
screen "eProC - 08 Descargador" 1280x768, template "Template"
   Button "Botón_4" at 220,383 size 93x33; TextOff 'Avance'
      on Press: SetTag("DB_OP.RC2", 70); SetBit("DB_OP.OP_SELMANU2")
      Visibility <- "MANU"
      Appearance <- "DB_OP.RC2"
   Button "Botón_5" at 220,421 size 93x33; TextOff 'Retroceso'
      on Press: SetTag("DB_OP.RC2", 71); SetBit("DB_OP.OP_SELMANU2")
      Visibility <- "MANU"
      Appearance <- "DB_OP.RC2"
   TextField "Campo de texto_5" at 229,340 size 85x23; Text 'Descargador'
      Visibility <- "MANU"
   Rectangle "Rectángulo_1" at 204,336 size 131x136
      Visibility <- "MANU"
   GraphicIOField "Campo ES gráfico_7" at 384,79 size 557x426; PictureList "Grupo 3 - Descargador"
      ProcessValue <- "Alarma_Descargador"
   Polygon "Polígono_4" at 443,271 size 39x59
      Visibility <- "Descargador-PiezaPresente"
   Polygon "Polígono_3" at 442,238 size 206x167
      Visibility <- "Descargador-PiezaPresente"
   Circle "Cercle_3" at 740,408 size 12x12
      Appearance <- "31S3"
   Circle "Cercle_4" at 693,373 size 12x12
      Appearance <- "31S8"
   Circle "Cercle_5" at 488,408 size 12x12
      Appearance <- "26S2"
   TextField "Campo de texto_1" at 890,544 size 173x22; Text '31S3 - Descargador Atrás'
   TextField "Campo de texto_2" at 557,516 size 195x22; Text '31S2 - Descargador Adelante'
   TextField "Campo de texto_3" at 818,279 size 193x22; Text '31S8 - Pieza en Descargador'
   Circle "Cercle_6" at 464,388 size 12x12
      Appearance <- "36S12"
   TextField "Campo de texto_4" at 534,549 size 294x22; Text '36S12 - Descargador en Posición Intermedia'
   Polygon "Polígono_2" at 450,217 size 81x72
      Visibility <- "Descargador-PiezaPresente"
   Polygon "Polígono_5" at 506,64 size 228x201
      Visibility <- "Descargador-PiezaPresente"
   Polygon "Polígono_1" at 543,118 size 206x170
      Visibility <- "Descargador-PiezaPresente"
   Polygon "Polígono_7" at 631,109 size 118x70
      Visibility <- "Descargador-PiezaPresente"
   Polygon "Polígono_8" at 625,64 size 112x67
      Visibility <- "Descargador-PiezaPresente"
   Rectangle "Rectángulo_2" at 204,336 size 131x32
      Visibility <- "MANU"
   Button "Template_Plantilla_Botón_3" at 1,688 size 130x29; TextOff 'DESCARGADOR'
   Button "Plantilla_Botón_1" at 1,715 size 130x53; TextOff 'PRINCIPAL'
      on Click: ActivateScreen("eProC - Principal", 0)
   Button "Template_Plantilla_Bouton_2" at 1085,715 size 193x53; TextOff 'ALARMAS / DEFAUT'
      on Press: ActivateScreen("eProC - Alarmas", 0)
      Visibility <- "DB_OP.P_DEFAUT"

screen "Gesión de Usuarios" 1280x768, template "Template"
   UserView "Visor de usuarios_1" at 28,48 size 1215x366
   Button "Botón_1" at 1059,488 size 176x56; TextOff 'Cerrar Sesión'
      on Activate: function_f23ef4c9()
   Button "Template_Plantilla_Botón_2" at 573,715 size 70x53; TextOff 'Text'; PictureOn "Usuario"; PictureOff "Usuario"; Authorization "Nivel 2"
      on Activate: ActivateScreen("Gesión de Usuarios", 0)
   Button "Template_Plantilla_Bouton_2" at 1085,715 size 193x53; TextOff 'ALARMAS / DEFAUT'
      on Press: ActivateScreen("eProC - Alarmas", 0)
      Visibility <- "DB_OP.P_DEFAUT"

screen "eProC - Historal" 1280x768, template "Template"
   AlarmView "Visor de avisos_1" at 29,48 size 1218x605; AlarmLog "Fichero_de_avisos_1"
   Button "Template_Plantilla_Botón_3" at 1085,688 size 193x29; TextOff 'HISTORIAL'
   Button "Template_Plantilla_Bouton_0" at 1085,715 size 193x53; TextOff 'ALARMAS / DEFAUT'
      on Press: ActivateScreen("eProC - Alarmas", 0)
   Button "Template_Plantilla_Bouton_2" at 1085,715 size 193x53; TextOff 'ALARMAS / DEFAUT'
      on Press: ActivateScreen("eProC - Alarmas", 0)
      Visibility <- "DB_OP.P_DEFAUT"

screen "eProC - Diagnóstico" 1280x768, template "Template"
   SysDiagControl "Sistema Visor de diagnóstico_1" at 16,30 size 1246x670; InfoArea_RootNodeText 'PLC Roll Forming / Installation'; NavigationPath_RootText 'Diagnóstico de Hardware / Vue d'ensemble du diagnostic'; NavigationpathDiagbufferText 'Búfer de diagnóstico / Vue du tampon de diagnostic'

screen "eProC - Estampado Alm 1" 1280x768, template "Template"
   TextField "Campo de texto_14" at 18,45 size 97x28; Text 'Almacén 1'
   TextField "Campo de texto_2" at 283,429 size 97x22; Text 'Herramienta 2'
   TextField "Campo de texto_3" at 283,157 size 97x22; Text 'Herramienta 1'
   TextField "Campo de texto_1" at 733,81 size 25x28; Text 'F1'
   TextField "Campo de texto_4" at 573,81 size 25x28; Text 'F3'
   TextField "Campo de texto_5" at 733,338 size 25x28; Text 'F2'
   TextField "Campo de texto_6" at 573,338 size 25x28; Text 'F4'
   TextField "Campo de texto_7" at 468,652 size 324x28; Text 'Resolución Incremento/Decremento'
   Button "Botón_1" at 754,150 size 40x40; TextOff 'Text'; PictureOff "outline_arrow_forward_ios_white_18dp"
      on Click: SetTag("PL_Dec_F_A1", 1)
   Button "Botón_2" at 698,150 size 40x40; TextOff 'Text'; PictureOff "outline_arrow_back_ios_white_18dp"
      on Click: SetTag("PL_Inc_F_A1", 1)
   Button "Botón_3" at 594,150 size 40x40; TextOff 'Text'; PictureOff "outline_arrow_forward_ios_white_18dp"
      on Click: SetTag("PL_Dec_F_A1", 3)
   Button "Botón_4" at 538,150 size 40x40; TextOff 'Text'; PictureOff "outline_arrow_back_ios_white_18dp"
      on Click: SetTag("PL_Inc_F_A1", 3)
   Button "Botón_5" at 754,406 size 40x40; TextOff 'Text'; PictureOff "outline_arrow_forward_ios_white_18dp"
      on Click: SetTag("PL_Dec_F_A1", 2)
   Button "Botón_6" at 698,406 size 40x40; TextOff 'Text'; PictureOff "outline_arrow_back_ios_white_18dp"
      on Click: SetTag("PL_Inc_F_A1", 2)
   Button "Botón_7" at 594,406 size 40x40; TextOff 'Text'; PictureOff "outline_arrow_forward_ios_white_18dp"
      on Click: SetTag("PL_Dec_F_A1", 4)
   Button "Botón_8" at 538,406 size 40x40; TextOff 'Text'; PictureOff "outline_arrow_back_ios_white_18dp"
      on Click: SetTag("PL_Inc_F_A1", 4)
   GraphicView "Visor de gráficos_7" at 263,452 size 138x75; Picture "F1-3 EMR2"
   GraphicView "Visor de gráficos_8" at 263,517 size 138x75; Picture "F2-4 EMR2"
   GraphicView "Visor de gráficos_2" at 263,180 size 138x75; Picture "EMR2"
   GraphicView "Visor de gráficos_3" at 263,245 size 138x75; Picture "F1-3 EMR2"
   IOField "Campo ES_1" at 698,109 size 96x32; FormatPattern s999999
      ProcessValue <- "Almacén 1\PAlmacén.F1"
   IOField "Campo ES_2" at 536,109 size 96x32; FormatPattern s999999
      ProcessValue <- "Almacén 1\PAlmacén.F3"
   IOField "Campo ES_3" at 698,366 size 96x32; FormatPattern s999999
      ProcessValue <- "Almacén 1\PAlmacén.F2"
   IOField "Campo ES_4" at 536,366 size 96x32; FormatPattern s999999
      ProcessValue <- "Almacén 1\PAlmacén.F4"
   IOField "Campo ES_5" at 787,653 size 96x32; FormatPattern 999999
      ProcessValue <- "PL_Resoluc_INCDECF"
   IOField "Champ E/S_1" at 122,48 size 410x24; FormatPattern ????????????????????
      ProcessValue <- "Almacén 1\PAlmacén.Nombre"

screen "eProC - Estampado Alm 2" 1280x768, template "Template"
   TextField "Campo de texto_14" at 18,45 size 97x28; Text 'Almacén 2'
   TextField "Campo de texto_2" at 283,429 size 97x22; Text 'Herramienta 2'
   TextField "Campo de texto_3" at 283,157 size 97x22; Text 'Herramienta 1'
   TextField "Campo de texto_1" at 733,81 size 25x28; Text 'F1'
   TextField "Campo de texto_4" at 572,81 size 25x28; Text 'F3'
   TextField "Campo de texto_5" at 733,338 size 25x28; Text 'F2'
   TextField "Campo de texto_6" at 572,338 size 25x28; Text 'F4'
   TextField "Campo de texto_7" at 468,652 size 324x28; Text 'Resolución Incremento/Decremento'
   Button "Botón_1" at 754,150 size 40x40; TextOff 'Text'; PictureOff "outline_arrow_forward_ios_white_18dp"
      on Click: SetTag("PL_Dec_F_A2", 1)
   Button "Botón_2" at 698,150 size 40x40; TextOff 'Text'; PictureOff "outline_arrow_back_ios_white_18dp"
      on Click: SetTag("PL_Inc_F_A2", 1)
   Button "Botón_3" at 593,150 size 40x40; TextOff 'Text'; PictureOff "outline_arrow_forward_ios_white_18dp"
      on Click: SetTag("PL_Dec_F_A2", 3)
   Button "Botón_4" at 537,150 size 40x40; TextOff 'Text'; PictureOff "outline_arrow_back_ios_white_18dp"
      on Click: SetTag("PL_Inc_F_A2", 3)
   Button "Botón_5" at 754,406 size 40x40; TextOff 'Text'; PictureOff "outline_arrow_forward_ios_white_18dp"
      on Click: SetTag("PL_Dec_F_A2", 2)
   Button "Botón_6" at 698,406 size 40x40; TextOff 'Text'; PictureOff "outline_arrow_back_ios_white_18dp"
      on Click: SetTag("PL_Inc_F_A2", 2)
   Button "Botón_7" at 593,406 size 40x40; TextOff 'Text'; PictureOff "outline_arrow_forward_ios_white_18dp"
      on Click: SetTag("PL_Dec_F_A2", 4)
   Button "Botón_8" at 537,406 size 40x40; TextOff 'Text'; PictureOff "outline_arrow_back_ios_white_18dp"
      on Click: SetTag("PL_Inc_F_A2", 4)
   GraphicView "Visor de gráficos_7" at 263,452 size 138x75; Picture "F1-3 EMR2"
   GraphicView "Visor de gráficos_8" at 263,517 size 138x75; Picture "F2-4 EMR2"
   GraphicView "Visor de gráficos_2" at 263,180 size 138x75; Picture "EMR2"
   GraphicView "Visor de gráficos_3" at 263,245 size 138x75; Picture "F1-3 EMR2"
   IOField "Campo ES_1" at 698,109 size 96x32; FormatPattern s999999
      ProcessValue <- "Almacén 2\PAlmacén.F1"
   IOField "Campo ES_2" at 535,109 size 96x32; FormatPattern s999999
      ProcessValue <- "Almacén 2\PAlmacén.F3"
   IOField "Campo ES_3" at 698,366 size 96x32; FormatPattern s999999
      ProcessValue <- "Almacén 2\PAlmacén.F2"
   IOField "Campo ES_4" at 535,366 size 96x32; FormatPattern s999999
      ProcessValue <- "Almacén 2\PAlmacén.F4"
   IOField "Campo ES_5" at 787,653 size 96x32; FormatPattern 999999
      ProcessValue <- "PL_Resoluc_INCDECF"
   IOField "Champ E/S_1" at 122,48 size 410x24; FormatPattern ????????????????????
      ProcessValue <- "Almacén 2\PAlmacén.Nombre"

screen "eProC - Plegado Alm 1" 1280x768, template "Template"
   TextField "Campo de texto_14" at 18,45 size 97x28; Text 'Almacén 1'
   TextField "Campo de texto_1" at 511,201 size 54x28; Text 'PL1-2'
   TextField "Campo de texto_4" at 773,201 size 54x28; Text 'PL2-2'
   TextField "Campo de texto_7" at 468,652 size 324x28; Text 'Resolución Incremento/Decremento'
   TextField "Campo de texto_2" at 1173,201 size 54x28; Text 'PL2-1'
   TextField "Campo de texto_3" at 110,201 size 54x28; Text 'PL1-1'
   IOField "Champ E/S_1" at 122,48 size 410x24; FormatPattern ????????????????????
      ProcessValue <- "Almacén 1\PAlmacén.Nombre"
   Button "Botón_1" at 543,270 size 40x40; TextOff 'Text'; PictureOff "outline_arrow_forward_ios_white_18dp"
      on Click: SetTag("PL_Dec_PL_A1", 2)
   Button "Botón_2" at 487,270 size 40x40; TextOff 'Text'; PictureOff "outline_arrow_back_ios_white_18dp"
      on Click: SetTag("PL_Inc_PL_A1", 2)
   Button "Botón_3" at 805,270 size 40x40; TextOff 'Text'; PictureOff "outline_arrow_forward_ios_white_18dp"
      on Click: SetTag("PL_Inc_PL_A1", 4)
   Button "Botón_4" at 749,270 size 40x40; TextOff 'Text'; PictureOff "outline_arrow_back_ios_white_18dp"
      on Click: SetTag("PL_Dec_PL_A1", 4)
   IOField "Campo ES_1" at 487,229 size 96x32; FormatPattern s999999
      ProcessValue <- "Almacén 1\PAlmacén.PL1_2"
   IOField "Campo ES_2" at 747,229 size 96x32; FormatPattern s999999
      ProcessValue <- "Almacén 1\PAlmacén.PL2_2"
   IOField "Campo ES_5" at 787,653 size 96x32; FormatPattern 999999
      ProcessValue <- "PL_Resoluc_INCDECPL"
   Button "Botón_9" at 1205,270 size 40x40; TextOff 'Text'; PictureOff "outline_arrow_forward_ios_white_18dp"
      on Click: SetTag("PL_Inc_PL_A1", 3)
   Button "Botón_10" at 1149,270 size 40x40; TextOff 'Text'; PictureOff "outline_arrow_back_ios_white_18dp"
      on Click: SetTag("PL_Dec_PL_A1", 3)
   IOField "Campo ES_6" at 1147,229 size 96x32; FormatPattern s999999
      ProcessValue <- "Almacén 1\PAlmacén.PL2_1"
   Button "Botón_11" at 142,270 size 40x40; TextOff 'Text'; PictureOff "outline_arrow_forward_ios_white_18dp"
      on Click: SetTag("PL_Dec_PL_A1", 1)
   Button "Botón_12" at 86,270 size 40x40; TextOff 'Text'; PictureOff "outline_arrow_back_ios_white_18dp"
      on Click: SetTag("PL_Inc_PL_A1", 1)
   IOField "Campo ES_7" at 86,229 size 96x32; FormatPattern s999999
      ProcessValue <- "Almacén 1\PAlmacén.PL1_1"

screen "eProC - Plegado Alm 2" 1280x768, template "Template"
   TextField "Campo de texto_14" at 18,45 size 97x28; Text 'Almacén 2'
   TextField "Campo de texto_1" at 511,201 size 54x28; Text 'PL1-2'
   TextField "Campo de texto_4" at 773,201 size 54x28; Text 'PL2-2'
   TextField "Campo de texto_7" at 468,652 size 324x28; Text 'Resolución Incremento/Decremento'
   TextField "Campo de texto_2" at 1173,201 size 54x28; Text 'PL2-1'
   TextField "Campo de texto_3" at 110,201 size 54x28; Text 'PL1-1'
   IOField "Champ E/S_1" at 122,48 size 410x24; FormatPattern ????????????????????
      ProcessValue <- "Almacén 2\PAlmacén.Nombre"
   Button "Botón_1" at 543,270 size 40x40; TextOff 'Text'; PictureOff "outline_arrow_forward_ios_white_18dp"
      on Click: SetTag("PL_Dec_PL_A2", 2)
   Button "Botón_2" at 487,270 size 40x40; TextOff 'Text'; PictureOff "outline_arrow_back_ios_white_18dp"
      on Click: SetTag("PL_Inc_PL_A2", 2)
   Button "Botón_3" at 805,270 size 40x40; TextOff 'Text'; PictureOff "outline_arrow_forward_ios_white_18dp"
      on Click: SetTag("PL_Inc_PL_A2", 4)
   Button "Botón_4" at 749,270 size 40x40; TextOff 'Text'; PictureOff "outline_arrow_back_ios_white_18dp"
      on Click: SetTag("PL_Dec_PL_A2", 4)
   IOField "Campo ES_1" at 487,229 size 96x32; FormatPattern s999999
      ProcessValue <- "Almacén 2\PAlmacén.PL1_2"
   IOField "Campo ES_2" at 747,229 size 96x32; FormatPattern s999999
      ProcessValue <- "Almacén 2\PAlmacén.PL2_2"
   IOField "Campo ES_5" at 787,653 size 96x32; FormatPattern 999999
      ProcessValue <- "PL_Resoluc_INCDECPL"
   Button "Botón_9" at 1205,270 size 40x40; TextOff 'Text'; PictureOff "outline_arrow_forward_ios_white_18dp"
      on Click: SetTag("PL_Inc_PL_A2", 3)
   Button "Botón_10" at 1149,270 size 40x40; TextOff 'Text'; PictureOff "outline_arrow_back_ios_white_18dp"
      on Click: SetTag("PL_Dec_PL_A2", 3)
   IOField "Campo ES_6" at 1147,229 size 96x32; FormatPattern s999999
      ProcessValue <- "Almacén 2\PAlmacén.PL2_1"
   Button "Botón_11" at 142,270 size 40x40; TextOff 'Text'; PictureOff "outline_arrow_forward_ios_white_18dp"
      on Click: SetTag("PL_Dec_PL_A2", 1)
   Button "Botón_12" at 86,270 size 40x40; TextOff 'Text'; PictureOff "outline_arrow_back_ios_white_18dp"
      on Click: SetTag("PL_Inc_PL_A2", 1)
   IOField "Campo ES_7" at 86,229 size 96x32; FormatPattern s999999
      ProcessValue <- "Almacén 2\PAlmacén.PL1_1"

screen "eProC - Principal" 1280x768, template "Template"
   Button "Button_4" at 186,452 size 74x115; TextOn 'Transfert en cours'; TextOff 'Transferencia / Transfert'
      on Press: ActivateScreen("eProC - 01 Araña", 0)
   Button "Button_3" at 130,516 size 74x51; TextOn 'Transfert en cours'; TextOff 'Transferencia / Transfert'
      on Press: ActivateScreen("eProC - 01 Araña", 0)
   Button "Button_5" at 242,468 size 82x67; TextOn 'Transfert en cours'; TextOff 'Transferencia / Transfert'
      on Press: ActivateScreen("eProC - 01 Araña", 0)
   Button "Button_8" at 322,486 size 90x51; TextOn 'Transfert en cours'; TextOff 'Transferencia / Transfert'
      on Press: ActivateScreen("eProC - 02 Rolos", 0)
   Button "Button_10" at 50,428 size 82x147; TextOn 'Transfert en cours'; TextOff 'Transferencia / Transfert'
      on Press: ActivateScreen("eProC - 00 Almacenes", 0)
   Button "Button_11" at 105,370 size 82x147; TextOn 'Transfert en cours'; TextOff 'Transferencia / Transfert'
      on Press: ActivateScreen("eProC - 00 Almacenes", 0)
   Button "Button_12" at 185,370 size 82x83; TextOn 'Transfert en cours'; TextOff 'Transferencia / Transfert'
      on Press: ActivateScreen("eProC - 00 Almacenes", 0)
   Button "Button_1" at 414,405 size 218x187; TextOn 'Transfert en cours'; TextOff 'Transferencia / Transfert'
      on Press: ActivateScreen("eProC - 03 Perfilador", 0)
   Button "Button_6" at 145,566 size 290x91; TextOn 'Transfert en cours'; TextOff 'Transferencia / Transfert'
      on Press: ActivateScreen("eProC - 02 Rolos", 0)
   Button "Button_7" at 257,534 size 178x35; TextOn 'Transfert en cours'; TextOff 'Transferencia / Transfert'
      on Press: ActivateScreen("eProC - 02 Rolos", 0)
   Button "Button_2" at 626,374 size 218x131; TextOn 'Transfert en cours'; TextOff 'Transferencia / Transfert'
      on Press: ActivateScreen("eProC - 10 - Estados F_HW", 0)
   Button "Button_9" at 746,374 size 162x35; TextOn 'Transfert en cours'; TextOff 'Transferencia / Transfert'
      on Press: ActivateScreen("eProC - 10 - Estados F_HW", 0)
   Button "Button_13" at 826,342 size 58x35; TextOn 'Transfert en cours'; TextOff 'Transferencia / Transfert'
      on Press: ActivateScreen("eProC - 10 - Estados F_HW", 0)
   Button "Button_14" at 666,286 size 161x89; TextOn 'Transfert en cours'; TextOff 'Transferencia / Transfert'
      on Press: ActivateScreen("eProC - 10 - Estados F_HW", 0)
   Button "Button_15" at 882,310 size 138x59; TextOn 'Transfert en cours'; TextOff 'Transferencia / Transfert'
      on Press: ActivateScreen("eProC - 10 - Estados F_HW", 0)
   Button "Button_16" at 914,302 size 98x123; TextOn 'Transfert en cours'; TextOff 'Transferencia / Transfert'
      on Press: ActivateScreen("eProC - 10 - Estados F_HW", 0)
   Button "Button_17" at 842,173 size 170x131; TextOn 'Transfert en cours'; TextOff 'Transferencia / Transfert'
      on Press: ActivateScreen("eProC - 09 - Estados PL_HW", 0)
   Button "Button_18" at 978,109 size 170x131; TextOn 'Transfert en cours'; TextOff 'Transferencia / Transfert'
      on Press: ActivateScreen("eProC - 09 - Estados PL_HW", 0)
   Button "Button_19" at 1018,245 size 210x179; TextOn 'Transfert en cours'; TextOff 'Transferencia / Transfert'
      on Press: ActivateScreen("eProC - 08 Descargador", 0)
   GraphicIOField "Campo ES gráfico_10" at 3,147 size 1272x557; PictureList "GeneralBase"
      ProcessValue <- "Alarma_General"
   GraphicIOField "Campo ES gráfico_7" at 827,154 size 309x174; PictureList "General - Plegadora"
      ProcessValue <- "Alarma_Plegador"
   GraphicIOField "Campo ES gráfico_2" at 58,421 size 219x150; PictureList "General - Almacén"
      ProcessValue <- "Alarma_Almacenes"
   GraphicIOField "Campo ES gráfico_8" at 758,313 size 77x78; PictureList "General - Formador"
      ProcessValue <- "Alarma_Formador"
   GraphicIOField "Campo ES gráfico_6" at 874,242 size 309x150; PictureList "General - Pinza"
      ProcessValue <- "Alarma_Pinza"
   GraphicIOField "Campo ES gráfico_5" at 610,339 size 293x150; PictureList "General - Cinta"
      ProcessValue <- "Alarma_Cinta"
   GraphicIOField "Campo ES gráfico_4" at 413,423 size 221x134; PictureList "General - Perfiladores"
      ProcessValue <- "Alarma_Perfiladores"
   GraphicIOField "Campo ES gráfico_3" at 148,495 size 285x158; PictureList "General - Rolos"
      ProcessValue <- "Alarma_Rolos"
   Polygon "Polígono_11" at 125,510 size 187x78
      Visibility <- "Araña\Araña.PresenciaPieza"
   Polygon "Polígono_1" at 423,444 size 190x70
      Visibility <- "Perfiladores\Perfilador.PresenciaPieza"
   Polygon "Polígono_3" at 184,523 size 186x78
      Visibility <- "Rolos\Rolos.PresenciaPieza"
   Polygon "Polígono_5" at 619,359 size 224x89
      Visibility <- "Cinta\Cinta.PresenciaPieza"
   GraphicIOField "Campo ES gráfico_1" at 46,380 size 300x302; PictureList "General - Araña"
      ProcessValue <- "Alarma_Araña"
   Polygon "Polígono_2" at 723,330 size 207x82
      Visibility <- "Pinza\Pinza.PresenciaPieza"
   Polygon "Polígono_10" at 871,196 size 265x104
      Visibility <- "Plegadora\Plegadora.PresenciaPieza"
   GraphicIOField "Campo ES gráfico_9" at 1016,197 size 141x246; PictureList "General - Descargador"
      ProcessValue <- "Alarma_Descargador"
   Polygon "Polígono_6" at 1065,227 size 66x79
      Visibility <- "Descargador-PiezaPresente"
   Polygon "Polígono_4" at 1026,266 size 35x54
      Visibility <- "Descargador-PiezaPresente"
   Polygon "Polígono_7" at 1044,306 size 19x15
      Visibility <- "Descargador-PiezaPresente"
   Polygon "Polígono_8" at 1044,228 size 58x75
      Visibility <- "Descargador-PiezaPresente"
   Polygon "Polígono_9" at 1062,293 size 17x17
      Visibility <- "Descargador-PiezaPresente"
   Polygon "Polígono_12" at 1063,309 size 17x8
      Visibility <- "Descargador-PiezaPresente"
   IOField "Campo ES_1" at 942,532 size 104x31; FormatPattern 9999.99; Unit  Segs.
      Visibility <- "eProC_Tiempos"
      ProcessValue <- "Tiempo_Heladera"
   IOField "Campo ES_2" at 1060,510 size 144x31; FormatPattern 9999.9; Unit  Helad/Hora
      ProcessValue <- "HxHoraInst"
      Visibility <- "eProC_Tiempos"
   TextField "Campo de texto_21" at 936,489 size 169x22; Text 'Tiempo entrega heladera'
      Visibility <- "eProC_Tiempos"
   IOField "Campo ES_3" at 1060,534 size 144x31; FormatPattern 9999.9; Unit  Helad/Hora
      ProcessValue <- "Tiempo_Heladera_1"
      Visibility <- "eProC_Tiempos"
   IOField "Campo ES_4" at 942,508 size 104x31; FormatPattern 9999.99; Unit  Segs.
      ProcessValue <- "Tiempo_Heladera_Parcial"
      Visibility <- "eProC_Tiempos"
   Button "Plantilla_Botón_1" at 1,715 size 130x53; TextOff 'PRINCIPAL'
      on Click: ActivateScreen("eProC - Principal", 0)
   IOField "Campo ES_5" at 109,69 size 64x39; FormatPattern 99999
      ProcessValue <- "ProD"
   Button "Botón_55" at 33,73 size 72x31; TextOff 'Reset'
      on Click: SetBit("Reset_ProD")
   TextField "Campo de texto_27" at 31,44 size 74x22; Text 'Producción'
   TextField "Campo de texto_28" at 353,44 size 73x22; Text 'Almacén 2'
   TextField "Campo de texto_29" at 211,44 size 73x22; Text 'Almacén 1'
   TextField "Campo de texto_30" at 394,78 size 21x22; Text 'de'
   TextField "Campo de texto_31" at 250,78 size 21x22; Text 'de'
   TextField "Campo de texto_33" at 578,44 size 43x22; Text 'Araña'
   TextField "Campo de texto_34" at 665,44 size 39x22; Text 'Rolos'
   TextField "Campo de texto_35" at 749,44 size 64x22; Text 'Perfilador'
   TextField "Campo de texto_38" at 939,44 size 38x22; Text 'Pinza'
   TextField "Campo de texto_39" at 1022,44 size 68x22; Text 'Plegadora'
   TextField "Campo de texto_113" at 857,44 size 37x22; Text 'Cinta'
   IOField "Champ E/S_11" at 276,76 size 48x26; FormatPattern 9999
      ProcessValue <- "DB_OP.M1_P_CPT"
   IOField "Champ E/S_12" at 211,73 size 45x31; FormatPattern 9999
      ProcessValue <- "DB_OP.M1_V_CPT"
   IOField "Champ E/S_13" at 420,76 size 47x26; FormatPattern 9999
      ProcessValue <- "DB_OP.M2_P_CPT"
   IOField "Champ E/S_14" at 355,73 size 45x31; FormatPattern 9999
      ProcessValue <- "DB_OP.M2_V_CPT"
   Button "Template_Plantilla_Bouton_2" at 1085,715 size 193x53; TextOff 'ALARMAS / DEFAUT'
      on Press: ActivateScreen("eProC - Alarmas", 0)
      Visibility <- "DB_OP.P_DEFAUT"
   IOField "Champ E/S_32" at 749,73 size 80x25; FormatPattern ????????????????????
      ProcessValue <- "Perfiladores\Perfilador.Nombre"
      Appearance <- "Perfiladores\Perfilador.PresenciaPieza"
   IOField "Champ E/S_33" at 665,73 size 80x25; FormatPattern ????????????????????
      ProcessValue <- "Rolos\Rolos.Nombre"
      Appearance <- "Rolos\Rolos.PresenciaPieza"
   IOField "Champ E/S_34" at 578,73 size 80x25; FormatPattern ????????????????????
      ProcessValue <- "Araña\Araña.Nombre"
      Appearance <- "Araña\Araña.PresenciaPieza"
   IOField "Champ E/S_35" at 857,73 size 80x25; FormatPattern ????????????????????
      ProcessValue <- "Cinta\Cinta.Nombre"
      Appearance <- "Cinta\Cinta.PresenciaPieza"
   IOField "Champ E/S_41" at 939,73 size 80x25; FormatPattern ????????????????????
      ProcessValue <- "Pinza\Pinza.Nombre"
      Appearance <- "Pinza\Pinza.PresenciaPieza"
   IOField "Champ E/S_42" at 1022,73 size 80x25; FormatPattern ????????????????????
      ProcessValue <- "Plegadora\Plegadora.Nombre"
      Appearance <- "Plegadora\Plegadora.PresenciaPieza"

screen "eProC - 09 - Estados PL" 1280x768, template "Template"
   Rectangle "Rectángulo_1" at 146,344 size 393x149
      Visibility <- "STOP_RUN"
   Button "Botón_2" at 352,429 size 144x40; TextOff 'Reset'
      on Click: SetBit("PL_Reset")
      Visibility <- "STOP_RUN"
   Button "Botón_1" at 192,429 size 144x40; TextOff 'Continuar'
      on Click: SetBit("PL_Continuar")
      Visibility <- "STOP_RUN"
   TextField "Campo de texto_17" at 165,356 size 351x73; Text 'Se ha detectado un reinicio del PLC. ¿Qué desea hacer con el ciclo de la Plegadora?'
      Visibility <- "STOP_RUN"
   IOField "Champ E/S_8" at 894,316 size 80x24; Authorization "Nivel 3"; FormatPattern 999; Unit  %
      ProcessValue <- "DB_OP.PL1_COD_VIT"
   IOField "Champ E/S_7" at 1077,316 size 80x24; Authorization "Nivel 3"; FormatPattern 999; Unit  %
      ProcessValue <- "DB_OP.PL2_COD_VIT"
   IOField "Champ E/S_4" at 894,240 size 91x29; Authorization "Nivel 2"; FormatPattern 9.9; Unit  
      ProcessValue <- "DB_OP.PL1_COD_COEF"
   IOField "Champ E/S_6" at 894,260 size 91x29; Authorization "Nivel 2"; FormatPattern s9999999; Unit  mm
      ProcessValue <- "DB_OP.PL1_COD_OFFSET"
   IOField "Champ E/S" at 1079,240 size 91x29; Authorization "Nivel 2"; FormatPattern 9.9; Unit  
      ProcessValue <- "DB_OP.PL2_COD_COEF"
   IOField "Champ E/S_2" at 1079,260 size 91x29; Authorization "Nivel 2"; FormatPattern s9999999; Unit  mm
      ProcessValue <- "DB_OP.PL2_COD_OFFSET"
   Button "Botón_4" at 815,462 size 94x45; TextOff 'Plegador 1'
      on Press: SetTag("Selec_Pleg", 1)
      Visibility <- "MANU"
      Appearance <- "Selec_Pleg"
   Button "Botón_9" at 918,462 size 94x45; TextOff 'Plegador 2'
      on Press: SetTag("Selec_Pleg", 2)
      Visibility <- "MANU"
      Appearance <- "Selec_Pleg"
   Button "Botón_10" at 711,462 size 94x45; TextOff 'General'
      on Press: SetTag("Selec_Pleg", 3)
      Visibility <- "MANU"
      Appearance <- "Selec_Pleg"
   SymbolicIOField "Campo ES simbólico_3" at 718,512 size 230x29; TextOn '1'; TextOff '0'; TextList "SelecciónPlegadora"
      Visibility <- "Selec_Pleg"
      ProcessValue <- "Selec_Pleg"
   Button "Botón_6" at 714,539 size 69x33; TextOff 'Subir'
      on Press: SetTag("DB_OP.RC2", 18); SetBit("DB_OP.OP_SELMANU2")
      Visibility <- "Selec_Pleg"
      Appearance <- "DB_OP.RC2"
   Button "Botón_7" at 714,576 size 69x33; TextOff 'Bajar'
      on Press: SetTag("DB_OP.RC2", 19); SetBit("DB_OP.OP_SELMANU2")
      Visibility <- "Selec_Pleg"
      Appearance <- "DB_OP.RC2"
   Button "Botón_8" at 790,539 size 77x33; TextOff 'Avance'
      on Press: SetTag("DB_OP.RC2", 61); SetBit("DB_OP.OP_SELMANU2")
      Visibility <- "Selec_Pleg"
      Appearance <- "DB_OP.RC2"
   Button "Botón_11" at 790,576 size 77x33; TextOff 'Retroceso'
      on Press: SetTag("DB_OP.RC2", 62); SetBit("DB_OP.OP_SELMANU2")
      Visibility <- "Selec_Pleg"
      Appearance <- "DB_OP.RC2"
   Button "Botón_12" at 873,539 size 69x33; TextOff 'Bloquear'
      on Press: SetTag("DB_OP.RC2", 10); SetBit("DB_OP.OP_SELMANU2")
      Visibility <- "Selec_Pleg"
      Appearance <- "DB_OP.RC2"
   Button "Botón_13" at 873,576 size 69x33; TextOff 'Desbloquear'
      on Press: SetTag("DB_OP.RC2", 11); SetBit("DB_OP.OP_SELMANU2")
      Visibility <- "Selec_Pleg"
      Appearance <- "DB_OP.RC2"
   Button "Botón_14" at 963,576 size 85x33; TextOff 'Bajar Prensa'
      on Press: SetTag("DB_OP.RC2", 12); SetBit("DB_OP.OP_SELMANU2")
      Visibility <- "Selec_Pleg"
      Appearance <- "DB_OP.RC2"
   Button "Botón_15" at 963,539 size 85x33; TextOff 'Subir Prensa'
      on Press: SetTag("DB_OP.RC2", 13); SetBit("DB_OP.OP_SELMANU2")
      Visibility <- "Selec_Pleg"
      Appearance <- "DB_OP.RC2"
   Button "Botón_17" at 1055,576 size 85x33; TextOff 'Bajar Ext 1'
      on Press: SetTag("DB_OP.RC2", 14); SetBit("DB_OP.OP_SELMANU2")
      Visibility <- "Selec_Pleg"
      Appearance <- "DB_OP.RC2"
   Button "Botón_18" at 1055,539 size 85x33; TextOff 'Subir Ext 1'
      on Press: SetTag("DB_OP.RC2", 15); SetBit("DB_OP.OP_SELMANU2")
      Visibility <- "Selec_Pleg"
      Appearance <- "DB_OP.RC2"
   Button "Botón_19" at 1146,576 size 85x33; TextOff 'Bajar Ext 2'
      on Press: SetTag("DB_OP.RC2", 16); SetBit("DB_OP.OP_SELMANU2")
      Visibility <- "Selec_Pleg"
      Appearance <- "DB_OP.RC2"
   Button "Botón_20" at 1146,539 size 85x33; TextOff 'Subir Ext 2'
      on Press: SetTag("DB_OP.RC2", 17); SetBit("DB_OP.OP_SELMANU2")
      Visibility <- "Selec_Pleg"
      Appearance <- "DB_OP.RC2"
   Polyline "Línea poligonal_5" at 1009,617 size 69x11
      Visibility <- "Selec_Pleg"
   TextField "Campo de texto_19" at 1081,618 size 40x18; Text 'Prensa'
      Visibility <- "Selec_Pleg"
   Polyline "Línea poligonal_6" at 1124,617 size 69x11
      Visibility <- "Selec_Pleg"
   Button "Botón_21" at 714,539 size 69x33; TextOff 'Subir'
      on Press: SetTag("DB_OP.RC2", 28); SetBit("DB_OP.OP_SELMANU2")
      Visibility <- "Selec_Pleg"
      Appearance <- "DB_OP.RC2"
   Button "Botón_22" at 714,576 size 69x33; TextOff 'Bajar'
      on Press: SetTag("DB_OP.RC2", 29); SetBit("DB_OP.OP_SELMANU2")
      Visibility <- "Selec_Pleg"
      Appearance <- "DB_OP.RC2"
   Button "Botón_23" at 790,539 size 77x33; TextOff 'Avance'
      on Press: SetTag("DB_OP.RC2", 65); SetBit("DB_OP.OP_SELMANU2")
      Visibility <- "Selec_Pleg"
      Appearance <- "DB_OP.RC2"
   Button "Botón_24" at 790,576 size 77x33; TextOff 'Retroceso'
      on Press: SetTag("DB_OP.RC2", 66); SetBit("DB_OP.OP_SELMANU2")
      Visibility <- "Selec_Pleg"
      Appearance <- "DB_OP.RC2"
   Button "Botón_25" at 873,539 size 69x33; TextOff 'Bloquear'
      on Press: SetTag("DB_OP.RC2", 20); SetBit("DB_OP.OP_SELMANU2")
      Visibility <- "Selec_Pleg"
      Appearance <- "DB_OP.RC2"
   Button "Botón_26" at 873,576 size 69x33; TextOff 'Desbloquear'
      on Press: SetTag("DB_OP.RC2", 21); SetBit("DB_OP.OP_SELMANU2")
      Visibility <- "Selec_Pleg"
      Appearance <- "DB_OP.RC2"
   Button "Botón_27" at 963,576 size 85x33; TextOff 'Bajar Prensa'
      on Press: SetTag("DB_OP.RC2", 22); SetBit("DB_OP.OP_SELMANU2")
      Visibility <- "Selec_Pleg"
      Appearance <- "DB_OP.RC2"
   Button "Botón_28" at 963,539 size 85x33; TextOff 'Subir Prensa'
      on Press: SetTag("DB_OP.RC2", 23); SetBit("DB_OP.OP_SELMANU2")
      Visibility <- "Selec_Pleg"
      Appearance <- "DB_OP.RC2"
   Button "Botón_29" at 1055,576 size 85x33; TextOff 'Bajar Ext 1'
      on Press: SetTag("DB_OP.RC2", 24); SetBit("DB_OP.OP_SELMANU2")
      Visibility <- "Selec_Pleg"
      Appearance <- "DB_OP.RC2"
   Button "Botón_30" at 1055,539 size 85x33; TextOff 'Subir Ext 1'
      on Press: SetTag("DB_OP.RC2", 25); SetBit("DB_OP.OP_SELMANU2")
      Visibility <- "Selec_Pleg"
      Appearance <- "DB_OP.RC2"
   Button "Botón_31" at 1146,576 size 85x33; TextOff 'Bajar Ext 2'
      on Press: SetTag("DB_OP.RC2", 26); SetBit("DB_OP.OP_SELMANU2")
      Visibility <- "Selec_Pleg"
      Appearance <- "DB_OP.RC2"
   Button "Botón_32" at 1146,539 size 85x33; TextOff 'Subir Ext 2'
      on Press: SetTag("DB_OP.RC2", 27); SetBit("DB_OP.OP_SELMANU2")
      Visibility <- "Selec_Pleg"
      Appearance <- "DB_OP.RC2"
   Polyline "Línea poligonal_3" at 1009,617 size 69x11
      Visibility <- "Selec_Pleg"
   TextField "Campo de texto_20" at 1081,618 size 40x18; Text 'Prensa'
      Visibility <- "Selec_Pleg"
   Polyline "Línea poligonal_4" at 1124,617 size 69x11
      Visibility <- "Selec_Pleg"
   Button "Botón_33" at 714,539 size 69x33; TextOff 'Subir'
      on Press: SetTag("DB_OP.RC2", 4); SetBit("DB_OP.OP_SELMANU2")
      Visibility <- "Selec_Pleg"
      Appearance <- "DB_OP.RC2"
   Button "Botón_34" at 714,576 size 69x33; TextOff 'Bajar'
      on Press: SetTag("DB_OP.RC2", 3); SetBit("DB_OP.OP_SELMANU2")
      Visibility <- "Selec_Pleg"
      Appearance <- "DB_OP.RC2"
   Button "Botón_35" at 790,539 size 77x33; TextOff 'Avance'
      on Press: SetTag("DB_OP.RC2", 1); SetBit("DB_OP.OP_SELMANU2")
      Visibility <- "Selec_Pleg"
      Appearance <- "DB_OP.RC2"
   Button "Botón_36" at 790,576 size 77x33; TextOff 'Retroceso'
      on Press: SetTag("DB_OP.RC2", 2); SetBit("DB_OP.OP_SELMANU2")
      Visibility <- "Selec_Pleg"
      Appearance <- "DB_OP.RC2"
   Button "Botón_37" at 873,539 size 69x33; TextOff 'Abrir'
      on Press: SetTag("DB_OP.RC2", 5); SetBit("DB_OP.OP_SELMANU2")
      Visibility <- "Selec_Pleg"
      Appearance <- "DB_OP.RC2"
   Button "Botón_38" at 873,576 size 69x33; TextOff 'Cerrar'
      on Press: SetTag("DB_OP.RC2", 6); SetBit("DB_OP.OP_SELMANU2")
      Visibility <- "Selec_Pleg"
      Appearance <- "DB_OP.RC2"
   Button "Botón_39" at 963,539 size 85x33; TextOff 'Alineación X'
      on Press: SetTag("DB_OP.RC2", 7); SetBit("DB_OP.OP_SELMANU2")
      Visibility <- "Selec_Pleg"
      Appearance <- "DB_OP.RC2"
   Button "Botón_40" at 963,576 size 85x33; TextOff 'Alineación Y'
      on Press: SetTag("DB_OP.RC2", 8); SetBit("DB_OP.OP_SELMANU2")
      Visibility <- "Selec_Pleg"
      Appearance <- "DB_OP.RC2"
   Button "Botón_41" at 1055,539 size 85x33; TextOff 'Subir Cepillos'
      on Press: SetTag("DB_OP.RC2", 9); SetBit("DB_OP.OP_SELMANU2")
      Visibility <- "Selec_Pleg"
      Appearance <- "DB_OP.RC2"
   Polyline "Línea poligonal_1" at 747,617 size 61x11
      Visibility <- "Selec_Pleg"
   TextField "Campo de texto_21" at 809,618 size 43x18; Text 'Tenaza'
      Visibility <- "Selec_Pleg"
   Polyline "Línea poligonal_2" at 857,617 size 61x11
      Visibility <- "Selec_Pleg"
   TextField "Template_Plantilla_Campo de texto_2" at 696,442 size 568x216; Text 'Text'
      Visibility <- "MANU"
   TextField "Template_Plantilla_Campo de texto_1" at 696,439 size 568x3; Text 'Text'
   Circle "Círculo_2" at 78,143 size 450x450
      Appearance <- "PL_en_Ciclo"
   SymbolicIOField "Campo ES simbólico_1" at 109,310 size 387x69; TextOn '1'; TextOff '0'; TextList "Estados_PL"
      ProcessValue <- "PL_Estados"
   Polygon "Polígono_1" at 466,215 size 12x13
      Appearance <- "PL_en_Ciclo"
   Polygon "Polígono_2" at 520,333 size 8x12
      Appearance <- "PL_en_Ciclo"
   Polygon "Polígono_3" at 503,456 size 8x12
      Appearance <- "PL_en_Ciclo"
   Polygon "Polígono_4" at 401,559 size 14x10
      Appearance <- "PL_en_Ciclo"
   Polygon "Polígono_5" at 242,583 size 14x7
      Appearance <- "PL_en_Ciclo"
   Polygon "Polígono_6" at 124,503 size 10x13
      Appearance <- "PL_en_Ciclo"
   Polygon "Polígono_7" at 78,389 size 6x17
      Appearance <- "PL_en_Ciclo"
   Polygon "Polígono_8" at 94,269 size 7x14
      Appearance <- "PL_en_Ciclo"
   Polygon "Polígono_9" at 345,145 size 13x6
      Appearance <- "PL_en_Ciclo"
   Polygon "Polígono_10" at 186,169 size 12x9
      Appearance <- "PL_en_Ciclo"
   GraphicIOField "Campo ES gráfico_1" at 90,461 size 50x46; PictureList "Estado"
      ProcessValue <- "PL_S_11"
   GraphicIOField "Campo ES gráfico_2" at 55,345 size 50x46; PictureList "Estado"
      ProcessValue <- "PL_S_6"
   GraphicIOField "Campo ES gráfico_4" at 196,137 size 50x46; PictureList "Estado"
      ProcessValue <- "PL_S_1"
   GraphicIOField "Campo ES gráfico_5" at 196,555 size 50x46; PictureList "Estado"
      ProcessValue <- "PL_S_5"
   GraphicIOField "Campo ES gráfico_6" at 356,137 size 50x46; PictureList "Estado"
      ProcessValue <- "PL_S_2"
   GraphicIOField "Campo ES gráfico_7" at 356,554 size 50x46; PictureList "Estado"
      ProcessValue <- "PL_S_10"
   GraphicIOField "Campo ES gráfico_8" at 467,464 size 50x46; PictureList "Estado"
      ProcessValue <- "PL_S_4"
   GraphicIOField "Campo ES gráfico_9" at 466,226 size 50x46; PictureList "Estado"
      ProcessValue <- "PL_S_9"
   GraphicIOField "Campo ES gráfico_10" at 501,345 size 50x46; PictureList "Estado"
      ProcessValue <- "PL_S_3"
   SymbolicIOField "Campo ES simbólico_2" at 103,359 size 403x45; TextOn '1'; TextOff '0'; TextList "Transiciones_PL"
      ProcessValue <- "PL_Estados"
   Line "Línea_1" at 109,126 size 0x102
      Appearance <- "PL_en_Ciclo"
   Polygon "Polígono_11" at 106,213 size 7x15
      Appearance <- "PL_en_Ciclo"
   GraphicIOField "Campo ES gráfico_11" at 84,121 size 50x46; PictureList "Estado"
      ProcessValue <- "PL_S_0"
   GraphicIOField "Campo ES gráfico_3" at 86,226 size 50x46; PictureList "Estado"
      ProcessValue <- "PL_S_12"
   TextField "Campo de texto_1" at 31,36 size 300x29; Text 'Máquina de estados Plegadores'
   IOField "Campo ES_1" at 890,72 size 80x32; FormatPattern 9999999; Unit  mm
      ProcessValue <- "PosiciónEspera_PL1"
      Appearance <- "PL_Req_Pos_Espera"
   TextField "Campo de texto_2" at 695,75 size 183x25; Text 'Posición de Espera'
      Appearance <- "PL_En_Pos_Espera"
   IOField "Campo ES_2" at 890,96 size 80x32; FormatPattern 9999999; Unit  mm
      ProcessValue <- "PosiciónRecepción_PL1"
      Appearance <- "PL_Req_Pos_Recep"
   TextField "Campo de texto_3" at 695,99 size 183x25; Text 'Posición de Recepción'
      Appearance <- "PL_En_Pos_Recepción"
   IOField "Campo ES_3" at 890,120 size 80x32; FormatPattern 9999999; Unit  mm
      ProcessValue <- "PosiciónPlegado1_PL1"
      Appearance <- "PL_Req_Pos_Pleg1"
   TextField "Campo de texto_4" at 695,123 size 183x25; Text 'Posición de Plegado Patas'
      Appearance <- "PL_En_Pos_Pleg1"
   IOField "Campo ES_4" at 890,144 size 80x32; FormatPattern 9999999; Unit  mm
      ProcessValue <- "PosiciónPlegado2_PL1"
      Appearance <- "PL_Req_Pos_Pleg2"
   TextField "Campo de texto_5" at 695,147 size 183x25; Text 'Posición de Plegado Techo'
      Appearance <- "PL_En_Pos_Pleg2"
   IOField "Campo ES_5" at 890,168 size 80x32; FormatPattern 9999999; Unit  mm
      ProcessValue <- "PosiciónEntrega_PL1"
      Appearance <- "PL_Req_Pos_Entrega"
   TextField "Campo de texto_6" at 695,171 size 183x25; Text 'Posición de Entrega'
      Appearance <- "PL_En_Pos_Entrega"
   IOField "Campo ES_6" at 1073,72 size 80x32; FormatPattern 9999999; Unit  mm
      ProcessValue <- "PosiciónEspera_PL2"
      Appearance <- "PL_Req_Pos_Espera"
   IOField "Campo ES_7" at 1073,96 size 80x32; FormatPattern 9999999; Unit  mm
      ProcessValue <- "PosiciónRecepción_PL2"
      Appearance <- "PL_Req_Pos_Recep"
   IOField "Campo ES_8" at 1073,120 size 80x32; FormatPattern 9999999; Unit  mm
      ProcessValue <- "PosiciónPlegado1_PL2"
      Appearance <- "PL_Req_Pos_Pleg1"
   IOField "Campo ES_9" at 1073,144 size 80x32; FormatPattern 9999999; Unit  mm
      ProcessValue <- "PosiciónPlegado2_PL2"
      Appearance <- "PL_Req_Pos_Pleg2"
   IOField "Campo ES_10" at 1073,168 size 80x32; FormatPattern 9999999; Unit  mm
      ProcessValue <- "PosiciónEntrega_PL2"
      Appearance <- "PL_Req_Pos_Entrega"
   TextField "Campo de texto_9" at 687,218 size 191x25; Text 'Límite Máximo de Posición'
   IOField "Campo ES_11" at 890,215 size 80x32; FormatPattern 9999999; Unit  mm
      ProcessValue <- "PosiciónMáxima_PL"
   IOField "Campo ES_12" at 1073,215 size 80x32; FormatPattern 9999999; Unit  mm
      ProcessValue <- "PosiciónMáxima_PL"
   TextField "Campo de texto_10" at 687,194 size 191x25; Text 'Límite Mínimo de Posición'
   IOField "Campo ES_13" at 890,191 size 80x32; FormatPattern 9999999; Unit  mm
      ProcessValue <- "PosiciónMínima_PL"
   IOField "Campo ES_14" at 1073,191 size 80x32; FormatPattern 9999999; Unit  mm
      ProcessValue <- "PosiciónMínima_PL"
   TextField "Campo de texto_11" at 727,288 size 151x25; Text 'Posición Actual'
   IOField "Campo ES_15" at 890,289 size 128x24; FormatPattern 9999999; Unit  mm
      ProcessValue <- "PosiciónActual_PL1"
   IOField "Campo ES_16" at 1073,289 size 128x24; FormatPattern 9999999; Unit  mm
      ProcessValue <- "PosiciónActual_PL2"
   TextField "Campo de texto_23" at 1160,381 size 82x36; Text 'MOVIMIENTO SEGURO'
      Visibility <- "PL_MovimientoSeguro"
      Appearance <- "PL_MovimientoSeguro"
   TextField "Campo de texto_12" at 727,319 size 151x17; Text 'Setpoint Velocidad'
   TextField "Campo de texto_15" at 372,147 size 16x25; Text '2'
   TextField "Campo de texto_16" at 482,236 size 16x25; Text '9'
   TextField "Campo de texto_13" at 518,355 size 16x25; Text '3'
   TextField "Campo de texto_24" at 483,474 size 16x25; Text '4'
   TextField "Campo de texto_26" at 366,564 size 30x25; Text '10'
   TextField "Campo de texto_27" at 211,565 size 19x25; Text '5'
   TextField "Campo de texto_28" at 100,471 size 30x25; Text '11'
   TextField "Campo de texto_29" at 70,355 size 15x25; Text '6'
   TextField "Campo de texto_30" at 96,236 size 31x25; Text '12'
   TextField "Campo de texto_31" at 212,147 size 16x25; Text '1'
   TextField "Campo de texto_32" at 100,131 size 16x25; Text '0'
   GraphicIOField "Campo ES gráfico_14" at 777,393 size 28x28; PictureList "CheckBox"
      ProcessValue <- "PL_Cepillos_No"
   GraphicIOField "Campo ES gráfico_15" at 840,393 size 28x28; PictureList "CheckBox"
      ProcessValue <- "PL_Prensas_No"
   GraphicIOField "Campo ES gráfico_16" at 912,393 size 28x28; PictureList "CheckBox"
      ProcessValue <- "PL_Fijaciones_No"
   GraphicIOField "Campo ES gráfico_17" at 998,393 size 28x28; PictureList "CheckBox"
      ProcessValue <- "PL_Alineado_No"
   GraphicIOField "Campo ES gráfico_18" at 1086,393 size 28x28; PictureList "CheckBox"
      ProcessValue <- "PL_Plegado_No"
   GraphicIOField "Campo ES gráfico_12" at 777,393 size 28x28; PictureList "CheckBox"
      ProcessValue <- "PL_S_1"
   IOField "Campo ES_17" at 972,72 size 80x32; FormatPattern 9999999; Unit  mm
      ProcessValue <- "PosiciónEspera_PL1(Ant)"
   IOField "Campo ES_18" at 972,96 size 80x32; FormatPattern 9999999; Unit  mm
      ProcessValue <- "PosiciónRecepción_PL1(Ant)"
   IOField "Campo ES_19" at 972,120 size 80x32; FormatPattern 9999999; Unit  mm
      ProcessValue <- "PosiciónPlegado1_PL1(Ant)"
   IOField "Campo ES_20" at 972,144 size 80x32; FormatPattern 9999999; Unit  mm
      ProcessValue <- "PosiciónPlegado2_PL1(Ant)"
   IOField "Campo ES_21" at 972,168 size 80x32; FormatPattern 9999999; Unit  mm
      ProcessValue <- "PosiciónEntrega_PL1(Ant)"
   IOField "Campo ES_22" at 1155,72 size 80x32; FormatPattern 9999999; Unit  mm
      ProcessValue <- "PosiciónEspera_PL2(Ant)"
   IOField "Campo ES_23" at 1155,96 size 80x32; FormatPattern 9999999; Unit  mm
      ProcessValue <- "PosiciónRecepción_PL2(Ant)"
   IOField "Campo ES_24" at 1155,120 size 80x32; FormatPattern 9999999; Unit  mm
      ProcessValue <- "PosiciónPlegado1_PL2(Ant)"
   IOField "Campo ES_25" at 1155,144 size 80x32; FormatPattern 9999999; Unit  mm
      ProcessValue <- "PosiciónPlegado2_PL2(Ant)"
   IOField "Campo ES_26" at 1155,168 size 80x32; FormatPattern 9999999; Unit  mm
      ProcessValue <- "PosiciónEntrega_PL2(Ant)"
   TextField "Campo de texto_33" at 894,37 size 81x23; Text 'Plegador 1'
   TextField "Campo de texto_34" at 1074,37 size 81x23; Text 'Plegador 2'
   Button "Botón_3" at 48,569 size 40x40; TextOff 'Vista Condiciones'; PictureOff "Gráfico_8"
      on Click: ActivateScreen("eProC - 09 - Estados PL_Diag", 0)
   TextField "Campo de texto_36" at 758,368 size 55x25; Text 'Cepillos'
   TextField "Campo de texto_37" at 823,368 size 55x25; Text 'Prensas'
   TextField "Campo de texto_38" at 887,368 size 71x25; Text 'Fijaciones'
   TextField "Campo de texto_39" at 975,368 size 71x25; Text 'Alineadores'
   TextField "Campo de texto_40" at 1063,368 size 71x25; Text 'Plegadores'
   TextField "Template_Plantilla_Campo de texto_3" at 696,359 size 568x3; Text 'Text'
   TextField "Template_Plantilla_Campo de texto_4" at 696,67 size 568x3; Text 'Text'
   Button "Botón_42" at 48,625 size 40x40; TextOff 'Vista Condiciones'; PictureOff "Gráfico_7"
      on Click: ActivateScreen("eProC - 09 - Estados PL_HW", 0)
   TextField "Campo de texto_22" at 687,242 size 191x25; Text 'Escalador relación mecánica'
   TextField "Campo de texto_25" at 687,262 size 191x25; Text 'Offset mecánico'
   TextField "Campo de texto_7" at 249,678 size 130x18; Text 'DATOS PIEZA ACTUAL'
   TextField "Campo de texto_8" at 403,678 size 12x18; Text 'A'
   IOField "Champ E/S_24" at 414,675 size 53x25; FormatPattern 9999999
      ProcessValue <- "Plegadora\Plegadora.A"
      Appearance <- "Plegadora\Plegadora.PresenciaPieza"
   IOField "Champ E/S_25" at 483,675 size 53x25; FormatPattern 9999999
      ProcessValue <- "Plegadora\Plegadora.B"
      Appearance <- "Plegadora\Plegadora.PresenciaPieza"
   IOField "Champ E/S_26" at 554,675 size 53x24; FormatPattern 9999999
      ProcessValue <- "Plegadora\Plegadora.C"
      Appearance <- "Plegadora\Plegadora.PresenciaPieza"
   IOField "Champ E/S_27" at 629,675 size 53x25; FormatPattern 9999999
      ProcessValue <- "Plegadora\Plegadora.D"
      Appearance <- "Plegadora\Plegadora.PresenciaPieza"
   TextField "Campo de texto_14" at 472,678 size 11x18; Text 'B'
   TextField "Campo de texto_18" at 541,678 size 11x18; Text 'C'
   TextField "Campo de texto_35" at 616,678 size 12x18; Text 'D'
   Button "Botón_5" at 1224,27 size 40x37; TextOff 'Vista Condiciones'; PictureOff "Tool"; Authorization "Nivel 3"
      on Click: ActivateScreen("eProC - 11 Referencias F-PL", 0)
   TextField "Campo de texto_41" at 700,37 size 75x23; Text 'Plegadora'
   Button "Template_Plantilla_Bouton_2" at 1085,715 size 193x53; TextOff 'ALARMAS / DEFAUT'
      on Press: ActivateScreen("eProC - Alarmas", 0)
      Visibility <- "DB_OP.P_DEFAUT"
   TextField "Campo de texto_170" at 717,678 size 35x18; Text 'PL1-1'
   IOField "Champ E/S_162" at 752,675 size 51x25; FormatPattern s999999
      ProcessValue <- "Plegadora\Plegadora.PL1_1"
      Appearance <- "Plegadora\Plegadora.PresenciaPieza"
   IOField "Champ E/S_163" at 857,675 size 51x25; FormatPattern s999999
      ProcessValue <- "Plegadora\Plegadora.PL1_2"
      Appearance <- "Plegadora\Plegadora.PresenciaPieza"
   IOField "Champ E/S_164" at 962,675 size 51x24; FormatPattern s999999
      ProcessValue <- "Plegadora\Plegadora.PL2_1"
      Appearance <- "Plegadora\Plegadora.PresenciaPieza"
   IOField "Champ E/S_165" at 1060,675 size 51x25; FormatPattern s999999
      ProcessValue <- "Plegadora\Plegadora.PL2_2"
      Appearance <- "Plegadora\Plegadora.PresenciaPieza"
   TextField "Campo de texto_171" at 821,678 size 35x18; Text 'PL1-2'
   TextField "Campo de texto_172" at 925,678 size 35x18; Text 'PL2-1'
   TextField "Campo de texto_173" at 1023,678 size 35x18; Text 'PL2-2'

